      Visibility <- "504_Tank Grouping_DB2020_GROUP of TANK 3"
   Circle "Circle_23" at 1000,464 size 14x14
      Appearance <- "20_TANKS_IP_DATA_RIO_01_THIRD_TANK_BWT_LEVEL_HIHI"
   TextField "Text field_126" at 955,465 size 51x14; Text 'LS422-1S'
   Polyline "Polyline_7" at 921,458 size 123x259
      Visibility <- "504_Tank Grouping_DB2020_RUN TANK 3"
   TextField "Text field_10" at 950,618 size 74x20; Text 'Tank - 1S'
   Bar "Bar_9" at 790,459 size 122x258; MinimumValue 0; MaximumValue 100
      ProcessValue <- "20_TANKS_IP_DATA_RIO_02_FIRST_TANK_TANKS_PRESS"
   Button "Button_34" at 801,662 size 100x25; TextOff 'DISABLED'
      on Release: function_efd93a16("Tank 2S Status", 168, 315, -1, 0, 1)
      Visibility <- "504_Tank Grouping_DB2020_GROUP of TANK 5"
   Circle "Circle_22" at 868,465 size 14x14
      Appearance <- "20_TANKS_IP_DATA_RIO_02_SECOND_TANK_BWT_LEVEL_HIHI"
   TextField "Text field_127" at 823,466 size 51x14; Text 'LS422-2S'
   Polyline "Polyline_8" at 789,458 size 123x259
      Visibility <- "504_Tank Grouping_DB2020_RUN TANK 5"
   TextField "Text field_11" at 817,618 size 74x20; Text 'Tank - 2S'
   Bar "Bar_10" at 659,460 size 122x258; MinimumValue 0; MaximumValue 100
      ProcessValue <- "20_TANKS_IP_DATA_RIO_03_FIRST_TANK_TANKS_PRESS"
   Button "Button_38" at 669,663 size 100x25; TextOff 'DISABLED'
      on Release: function_efd93a16("Tank 3S Status", 168, 315, -1, 0, 1)
      Visibility <- "504_Tank Grouping_DB2020_GROUP of TANK 7"
   Circle "Circle_21" at 736,467 size 14x14
      Appearance <- "20_TANKS_IP_DATA_RIO_03_SECOND_TANK_BWT_LEVEL_HIHI"
   TextField "Text field_128" at 691,468 size 51x14; Text 'LS422-3S'
   Polyline "Polyline_9" at 658,458 size 123x259
      Visibility <- "504_Tank Grouping_DB2020_RUN TANK 7"
   TextField "Text field_12" at 690,618 size 74x20; Text 'Tank - 3S'
   Bar "Bar_11" at 526,459 size 122x258; MinimumValue 0; MaximumValue 100
      ProcessValue <- "20_TANKS_IP_DATA_RIO_04_FIRST_TANK_TANKS_PRESS"
   Button "Button_42" at 537,662 size 100x25; TextOff 'DISABLED'
      on Release: function_efd93a16("Tank 4S Status", 168, 315, -1, 2, 1)
      Visibility <- "504_Tank Grouping_DB2020_GROUP of TANK 9"
   Circle "Circle_19" at 604,466 size 14x14
      Appearance <- "20_TANKS_IP_DATA_RIO_04_SECOND_TANK_BWT_LEVEL_HIHI"
   TextField "Text field_129" at 559,467 size 51x14; Text 'LS422-4S'
   Polyline "Polyline_10" at 525,458 size 123x259
      Visibility <- "504_Tank Grouping_DB2020_RUN TANK 9"
   TextField "Text field_13" at 554,618 size 74x20; Text 'Tank - 4S'
   Bar "Bar_12" at 394,459 size 122x258; MinimumValue 0; MaximumValue 100
      ProcessValue <- "20_TANKS_IP_DATA_RIO_05_FIRST_TANK_TANKS_PRESS"
   Button "Button_46" at 405,662 size 100x25; TextOff 'DISABLED'
      on Release: function_efd93a16("Tank 5S Status", 168, 315, -1, 2, 1)
      Visibility <- "504_Tank Grouping_DB2020_GROUP of TANK 11"
   Circle "Circle_18" at 472,465 size 14x14
      Appearance <- "20_TANKS_IP_DATA_RIO_05_SECOND_TANK_BWT_LEVEL_HIHI"
   TextField "Text field_130" at 427,466 size 51x14; Text 'LS422-5S'
   Polyline "Polyline_11" at 393,458 size 123x259
      Visibility <- "504_Tank Grouping_DB2020_RUN TANK 11"
   TextField "Text field_18" at 424,618 size 74x20; Text 'Tank - 5S'
   Bar "Bar_13" at 262,460 size 122x258; MinimumValue 0; MaximumValue 100
      ProcessValue <- "20_TANKS_IP_DATA_RIO_06_FIRST_TANK_TANKS_PRESS"
   Button "Button_50" at 273,663 size 100x25; TextOff 'DISABLED'
      on Release: function_efd93a16("Tank 6S Status", 168, 315, -1, 2, 1)
      Visibility <- "504_Tank Grouping_DB2020_GROUP of TANK 13"
   Circle "Circle_17" at 340,467 size 14x14
      Appearance <- "20_TANKS_IP_DATA_RIO_06_SECOND_TANK_BWT_LEVEL_HIHI"
   TextField "Text field_131" at 295,468 size 51x14; Text 'LS422-6S'
   Polyline "Polyline_12" at 261,458 size 123x258
      Visibility <- "504_Tank Grouping_DB2020_RUN TANK 13"
   TextField "Text field_19" at 290,618 size 74x20; Text 'Tank - 6S'
   Bar "Bar_14" at 39,324 size 119x258; Unit %; MinimumValue 0; MaximumValue 100
      ProcessValue <- "20_TANKS_IP_DATA_RIO_07_FIRST_TANK_TANKS_PRESS"
   Circle "Circle_25" at 108,330 size 14x14
      Appearance <- "20_TANKS_IP_DATA_RIO_07_FIRST_TANK_BWT_LEVEL_HIHI"
   TextField "Text field_132" at 79,330 size 35x14; Text 'LS425'
   Polyline "Polyline_13" at 38,324 size 121x259
      Visibility <- "504_Tank Grouping_DB2020_RUN TANK 14"
   Button "Button_58" at 48,527 size 100x25; TextOff 'DISABLED'
      on Release: function_efd93a16("Tank AP Status", 168, 315, -1, 2, 1)
      Visibility <- "504_Tank Grouping_DB2020_GROUP of TANK 14"
   Button "HmiScreenItemData_6" at 1043,144 size 116x50; TextOn 'Back'; TextOff 'Tank Status'
      on Release: ActivateScreen("Balast Water Treatment Plant", 0)
   Button "Button_2" at 252,437 size 37x30; TextOff 'DB&B'
      on Release: function_efd93a16("Double Block & Bleed Valve Monitoring", 250, 250, -1, -1, 1)
      Appearance <- "10_DI_DATA_CV407_OPN"
   TextField "Text field_65" at 190,398 size 46x25; Text 'PGC'
   TextField "Text field_75" at 183,480 size 60x20; Text 'Disabled'
   TextField "Text field_76" at 183,480 size 60x20; Text 'Enabled'
      Visibility <- "10_DI_DATA_E_400_RUN"
   GraphicView "Graphic view_76" at 185,421 size 57x55; Picture "Graphic_251"
   Button "Button_6" at 179,402 size 70x105; TextOff 'Text'
      on Release: ActivateScreen("PGC System", 0)
   TextField "Text field_20" at 53,396 size 103x20; Text 'Aft PeakTank'
   GraphicView "Graphic view_108" at 4,683 size 96x48; Picture "Left Arow"
   Button "HmiScreenItemData_14" at 3,660 size 106x93; TextOn 'Back'; TextOff 'Text'
      on Press: ActivateScreen("Inert Gas Conditioning Plant", 0)
   IOField "I/O field_1" at 44,460 size 115x25; FormatPattern s999.9; Unit mBar
      ProcessValue <- "20_TANKS_IP_DATA_RIO_07_FIRST_TANK_TANKS_PRESS"
   IOField "I/O field_2" at 269,331 size 114x25; FormatPattern s999.9; Unit mBar
      ProcessValue <- "20_TANKS_IP_DATA_RIO_06_FIRST_TANK_TANKS_PRESS"
   IOField "I/O field_3" at 398,331 size 117x25; FormatPattern s999.9; Unit mBar
      ProcessValue <- "20_TANKS_IP_DATA_RIO_05_FIRST_TANK_TANKS_PRESS"
   IOField "I/O field_4" at 531,331 size 117x25; FormatPattern s999.9; Unit mBar
      ProcessValue <- "20_TANKS_IP_DATA_RIO_04_FIRST_TANK_TANKS_PRESS"
   IOField "I/O field_5" at 662,331 size 114x25; FormatPattern s999.9; Unit mBar
      ProcessValue <- "20_TANKS_IP_DATA_RIO_03_FIRST_TANK_TANKS_PRESS"
   IOField "I/O field_6" at 796,331 size 119x25; FormatPattern s999.9; Unit mBar
      ProcessValue <- "20_TANKS_IP_DATA_RIO_02_FIRST_TANK_TANKS_PRESS"
   IOField "I/O field_7" at 928,331 size 118x25; FormatPattern s999.9; Unit mBar
      ProcessValue <- "20_TANKS_IP_DATA_RIO_01_FIRST_TANK_TANKS_PRESS"
   IOField "I/O field_8" at 1103,459 size 119x25; FormatPattern s999.9; Unit mBar
      ProcessValue <- "20_TANKS_IP_DATA_RIO_01_FIRST_TANK_TANKS_PRESS"
   IOField "I/O field_9" at 928,555 size 118x25; FormatPattern s999.9; Unit mBar
      ProcessValue <- "20_TANKS_IP_DATA_RIO_01_FIRST_TANK_TANKS_PRESS"
   IOField "I/O field_10" at 796,556 size 118x25; FormatPattern s999.9; Unit mBar
      ProcessValue <- "20_TANKS_IP_DATA_RIO_02_FIRST_TANK_TANKS_PRESS"
   IOField "I/O field_11" at 664,558 size 116x25; FormatPattern s999.9; Unit mBar
      ProcessValue <- "20_TANKS_IP_DATA_RIO_03_FIRST_TANK_TANKS_PRESS"
   IOField "I/O field_12" at 530,557 size 117x25; FormatPattern s999.9; Unit mBar
      ProcessValue <- "20_TANKS_IP_DATA_RIO_04_FIRST_TANK_TANKS_PRESS"
   IOField "I/O field_13" at 400,558 size 114x25; FormatPattern s999.9; Unit mBar
      ProcessValue <- "20_TANKS_IP_DATA_RIO_05_FIRST_TANK_TANKS_PRESS"
   IOField "I/O field_14" at 268,559 size 116x25; FormatPattern s999.9; Unit mBar
      ProcessValue <- "20_TANKS_IP_DATA_RIO_06_FIRST_TANK_TANKS_PRESS"
   Button "Button_88" at 34,324 size 127x264; TextOff 'Text'
      on Release: function_efd93a16("Tank AP Status", 168, 315, -1, 0, 1)
      Appearance <- "504_Tank Grouping_DB2020_RUN TANK 14"
   Button "Button_86" at 259,458 size 126x260; TextOff 'Text'
      on Release: function_efd93a16("Tank 6S Status", 168, 315, -1, 0, 1)
      Appearance <- "504_Tank Grouping_DB2020_RUN TANK 13"
   Button "Button_79" at 391,457 size 126x262; TextOff 'Text'
      on Release: function_efd93a16("Tank 5S Status", 168, 315, -1, 0, 1)
      Appearance <- "504_Tank Grouping_DB2020_RUN TANK 11"
   Button "Button_77" at 523,457 size 126x262; TextOff 'Text'
      on Release: function_efd93a16("Tank 4S Status", 168, 315, -1, 0, 1)
      Appearance <- "504_Tank Grouping_DB2020_RUN TANK 9"
   Button "Button_74" at 657,457 size 126x262; TextOff 'Text'
      on Release: function_efd93a16("Tank 3S Status", 168, 315, -1, 0, 1)
      Appearance <- "504_Tank Grouping_DB2020_RUN TANK 7"
   Button "Button_70" at 788,457 size 126x262; TextOff 'Text'
      on Release: function_efd93a16("Tank 2S Status", 168, 315, -1, 0, 1)
      Appearance <- "504_Tank Grouping_DB2020_RUN TANK 5"
   Button "Button_66" at 921,457 size 126x261; TextOff 'Text'
      on Release: function_efd93a16("Tank 1S Status", 168, 315, -1, 0, 1)
      Appearance <- "504_Tank Grouping_DB2020_RUN TANK 3"
   Button "Button_61" at 1093,328 size 130x248; TextOff 'Text'
      on Release: function_efd93a16("Tank FP Status", 168, 315, -1, 0, 1)
      Appearance <- "504_Tank Grouping_DB2020_RUN TANK 1"
   Button "Button_62" at 919,205 size 126x242; TextOff 'Text'
      on Release: function_efd93a16("Tank 1P Status", 168, 315, -1, 0, 1)
      Appearance <- "504_Tank Grouping_DB2020_RUN TANK 2"
   Button "Button_68" at 789,202 size 126x246; TextOff 'Text'
      on Release: function_efd93a16("Tank 2P Status", 168, 315, -1, 0, 1)
      Appearance <- "504_Tank Grouping_DB2020_RUN TANK 4"
   Button "Button_72" at 654,205 size 126x242; TextOff 'Text'
      on Release: function_efd93a16("Tank 3P Status", 168, 315, -1, 0, 1)
      Appearance <- "504_Tank Grouping_DB2020_RUN TANK 6"
   Button "Button_76" at 524,205 size 126x243; TextOff 'Text'
      on Release: function_efd93a16("Tank 4P Status", 168, 315, -1, 0, 1)
      Appearance <- "504_Tank Grouping_DB2020_RUN TANK 8"
   Button "Button_78" at 392,206 size 126x241; TextOff 'Text'
      on Release: function_efd93a16("Tank 5P Status", 168, 315, -1, 0, 1)
      Appearance <- "504_Tank Grouping_DB2020_RUN TANK 10"
   Button "Button_84" at 259,204 size 126x244; TextOff 'Text'
      on Release: function_efd93a16("Tank 6P Status", 168, 315, -1, 0, 1)
      Appearance <- "504_Tank Grouping_DB2020_RUN TANK 12"
   Group "Group_5" at 664,46 size 45x27; FormatPattern 999
   Group "Group_1" at 711,46 size 50x27; FormatPattern 999; Unit h
   Group "Group_2" at 605,46 size 57x27; FormatPattern 999; Unit h
   Button "HmiScreenItemData_5" at 180,144 size 116x50; TextOn 'Back'; TextOff 'Tank Status'
      on Release: function_efd93a16("Tank Status", 400, 250, -1, -1, 1)
   Button "Button_10" at 14,93 size 153x55; TextOff 'Text'
      on Release: function_efd93a16("Salinity - Acceptance", 168, 315, -1, 0, 1)
      Visibility <- "2068_Sys_Status_Data_SAL_VALID"
   Button "Button_12" at 14,93 size 153x53; TextOff 'Text'
      on Release: function_efd93a16("Tank Times", 300, 200, -1, 0, 1)
      Visibility <- "2068_Sys_Status_Data_Times Visibil"
   Button "Button_59" at 298,44 size 240x30; TextOn 'TB3 Enabled'; TextOff 'BWT System Shutting Down'
      Visibility <- "2110_BTCS_CNTRL_DB_BTCS_STATE"
   Button "Button_60" at 299,44 size 240x30; TextOn 'TB3 Enabled'; TextOff 'BWT System Enabled'
      Visibility <- "2110_BTCS_CNTRL_DB_BTCS_STATE"
   IOField "I/O field_29" at 664,46 size 45x27; FormatPattern 99; Unit h
      ProcessValue <- "Sequence Times_DB_Treatment Timer_Hours Left"
      Visibility <- "2110_BTCS_CNTRL_DB_BTCS_STATE"
   IOField "I/O field_30" at 664,46 size 45x27; FormatPattern 99; Unit h
      ProcessValue <- "Sequence Times_DB_Pre-Dwell Timer_Hours Left"
      Visibility <- "2110_BTCS_CNTRL_DB_BTCS_STATE"
   IOField "I/O field_15" at 711,46 size 50x27; FormatPattern 99; Unit m
      ProcessValue <- "Sequence Times_DB_Treatment Timer_Minutes Left"
      Visibility <- "2110_BTCS_CNTRL_DB_BTCS_STATE"
   IOField "I/O field_16" at 711,46 size 50x27; FormatPattern 99; Unit m
      ProcessValue <- "Sequence Times_DB_Pre-Dwell Timer_Minutes Left"
      Visibility <- "2110_BTCS_CNTRL_DB_BTCS_STATE"
   IOField "I/O field_17" at 605,46 size 57x27; FormatPattern 999; Unit d
      ProcessValue <- "Sequence Times_DB_Treatment Timer_Days Left"
      Visibility <- "2110_BTCS_CNTRL_DB_BTCS_STATE"
   IOField "I/O field_18" at 605,46 size 57x27; FormatPattern 999; Unit d
      ProcessValue <- "Sequence Times_DB_Pre-Dwell Timer_Days Left"
      Visibility <- "2110_BTCS_CNTRL_DB_BTCS_STATE"

VB script "VoyageTimeInsufficient"
   If SmartTags("Voyage Time Invalid") Then
   	efd93a16-2665-4b85-bcb9-25eddcb7b6f4 Voyage Time Warning,275,250,$3$hmiOn$,$3$hmiTop$,$3$hmiMedium$
   ElseIf Not SmartTags("Voyage Time Invalid") Then
   	efd93a16-2665-4b85-bcb9-25eddcb7b6f4Voyage Time Warning,0,0,$3$hmiOff$,$3$hmiAnimationOff$,$3$hmiMedium$
   End If

VB script "TreatmentCycleCompleted"
   If SmartTags("Sequence Times_DB_Post-Dwell Timer_Q") Then
   	efd93a16-2665-4b85-bcb9-25eddcb7b6f4 Treatment Cycle Completed,275,250,$3$hmiOn$,$3$hmiBottom$,$3$hmiMedium$
   'ElseIf Not SmartTags("Treatment Runs Completed") Then
   '	ShowPopupScreen"Treatment Cycle Completed",0,0,hmiOff,hmiAnimationOff,hmiMedium
   End If

VB script "SD_Card_Overflow"
   If SmartTags("Logging SD Card Overflow") Then 
   	efd93a16-2665-4b85-bcb9-25eddcb7b6f4 SD Card overflow,275,250,$3$hmiOn$,$3$hmiBottom$,$3$hmiMedium$
   ElseIf Not SmartTags("Logging SD Card Overflow") Then
   	efd93a16-2665-4b85-bcb9-25eddcb7b6f4SD Card overflow,0,0,$3$hmiOff$,$3$hmiAnimationOff$,$3$hmiMedium$
   End If

VB script "Salinity_FreshWaterAlert"
   If SmartTags("2068_Sys_Status_Data_SAL_CNF_CHK") Then
   	efd93a16-2665-4b85-bcb9-25eddcb7b6f4 Salinity - Fresh Water Alert,789,316,$3$hmiOn$,$3$hmiBottom$,$3$hmiMedium$
   ElseIf Not SmartTags("2068_Sys_Status_Data_SAL_CNF_CHK") Then
   	efd93a16-2665-4b85-bcb9-25eddcb7b6f4Salinity - Fresh Water Alert,0,0,$3$hmiOff$,$3$hmiAnimationOff$,$3$hmiMedium$
   End If

VB script "TimeRemainingToTreatment"
   If SmartTags("Warn To Start IGG") Then
   	efd93a16-2665-4b85-bcb9-25eddcb7b6f4 Time Until Treatment Required, 400, 200, $3$hmiOn$, $3$hmiBottom$, $3$hmiMedium$
   	ElseIf Not SmartTags("Warn To Start IGG") Then
   efd93a16-2665-4b85-bcb9-25eddcb7b6f4 Time Until Treatment Required, 0, 0, $3$hmiOff$, $3$hmiOff$, $3$hmiMedium$
   End If

VB script "TreatmentRequired"
   If SmartTags("Warn To Start IGG-Last") Then
   	efd93a16-2665-4b85-bcb9-25eddcb7b6f4 Start Treatment, 400, 200, $3$hmiOn$, $3$hmiBottom$, $3$hmiMedium$
   	ElseIf Not SmartTags("Warn To Start IGG-Last") Then
   efd93a16-2665-4b85-bcb9-25eddcb7b6f4 Start Treatment, 0, 0, $3$hmiOff$, $3$hmiOff$, $3$hmiMedium$
   End If

VB script "PGCCommissioning"
   If SmartTags("PGC_COMMISSION_MODE_DB_Drive Popup") Then
   	efd93a16-2665-4b85-bcb9-25eddcb7b6f4 PGC Commissioning, 0, 0, $3$hmiOn$, $3$hmiBottom$, $3$hmiMedium$
   	ElseIf Not SmartTags("PGC_COMMISSION_MODE_DB_Drive Popup") Then
   efd93a16-2665-4b85-bcb9-25eddcb7b6f4 PGC Commissioning, 0, 0, $3$hmiOff$, $3$hmiOff$, $3$hmiMedium$
   End If

VB script "User_Change"
   f41c6f6c-971d-4734-9362-16d81ac70597 Current User
   e1ab61de-e5a2-437b-97c4-abda991a3a2e user_group
   
   'Tip:
   ' 1. Use the <CTRL+SPACE> or <CTRL+I> shortcut to open a list of all objects and functions
   ' 2. Write the code using the HMI Runtime object.
   '  Example: HmiRuntime.Screens("Screen_1").
   ' 3. Use the <CTRL+J> shortcut to create an object reference.
   'Write the code as of this position:

VB script "TreatmentdDailyChecks"
   If SmartTags("88_treatment_POP_UP") Then
   	efd93a16-2665-4b85-bcb9-25eddcb7b6f4 Treatment check / Daily Checks Completed,275,250,$3$hmiOn$,$3$hmiBottom$,$3$hmiMedium$
   End If

VB script "TitleUpdater"
   Dim title
   Set title = HmiRuntime.ActiveScreen.ScreenItems("Screen title")
   title.Text = HmiRuntime.ActiveScreen.ObjectName

VB script "BWT_Warning"
   If SmartTags("2068_Sys_Status_Data_Not BWT mode Warning") Then
   	efd93a16-2665-4b85-bcb9-25eddcb7b6f4 BWT Mode Warning,275,250,$3$hmiOn$,$3$hmiTop$,$3$hmiMedium$
   'ElseIf Not SmartTags("BWT Mode Warning") Then
   '	ShowPopupScreen"BWT Mode Warning",0,0,hmiOff,hmiAnimationOff,hmiMedium
   End If

VB script "Report_Test"
   f41c6f6c-971d-4734-9362-16d81ac70597 Current User
   e1ab61de-e5a2-437b-97c4-abda991a3a2e user_group
   
   
   'Tip:
   ' 1. Use the <CTRL+SPACE> or <CTRL+I> shortcut to open a list of all objects and functions
   ' 2. Write the code using the HMI Runtime object.
   '  Example: HmiRuntime.Screens("Screen_1").
   ' 3. Use the <CTRL+J> shortcut to create an object reference.
   'Write the code as of this position:

VB script "HeartBeatFunction"
   If SmartTags("IGG HMI HEART BEAT")=0 Then
   	b21d3eaf-4e31-425c-ad1a-ba4e4002cacc(IGG HMI HEART BEAT),1
   Else
   	b21d3eaf-4e31-425c-ad1a-ba4e4002cacc (IGG HMI HEART BEAT),0
   End If

VB script "HeartBeatHMI_Warning"
   Dim Warning, Tempos
   
   
   If SmartTags("HEART BEAT TRUE")=True Then
   	Warning=0 '"HEART BEAT TRUE"
   Else
   	Warning=1
   End If
   
   If Warning=0 Then
   	efd93a16-2665-4b85-bcb9-25eddcb7b6f4 Lost Comunication, 0, 0, $3$hmiOff$, $3$hmiOff$, $3$hmiMedium$
   Else
   	efd93a16-2665-4b85-bcb9-25eddcb7b6f4 Lost Comunication, 300, 100, $3$hmiOn$, $3$hmiBottom$, $3$hmiMedium$
   End If		
   
   	b21d3eaf-4e31-425c-ad1a-ba4e4002cacc SmartTags("HEART BEAT TRUE"),False

VB script "PGC_ProtectionWarning"
   If SmartTags("Setpoint Override_DB_Set Pressure") Then
   	efd93a16-2665-4b85-bcb9-25eddcb7b6f4 PGC Protection Warning,275,250,$3$hmiOn$,$3$hmiTop$,$3$hmiMedium$
   'ElseIf Not SmartTags("Setpoint Override_DB_Set Pressure") Then
   '	ShowPopupScreen"Setpoint Override_DB_Set Pressure",0,0,hmiOff,hmiAnimationOff,hmiMedium
   End If

VB script "ALARM_Present"
   If SmartTags("60_Alarm_Data_ALRM_PRSNT") Then
   	bec8f1e5-2ab1-45f6-ad91-1d37c469eb91 04 Alarm Log,0
   End If
   
   'If Not SmartTags("60_Alarm_Data_ALRM_PRSNT") Then
   '	ActivateScreen "01 Home",0
   'End If
   
   
   
   
   
   
   
   
   
   'Tip:
   ' 1. Use the <CTRL+SPACE> or <CTRL+I> shortcut to open a list of all objects and functions
   ' 2. Write the code using the HMI Runtime object.
   '  Example: HmiRuntime.Screens("Screen_1").
   ' 3. Use the <CTRL+J> shortcut to create an object reference.
   'Write the code as of this position:

VB script "TreatmentRequired_GCU"
   If SmartTags("Warn To Start GCU-Last") Then
   	efd93a16-2665-4b85-bcb9-25eddcb7b6f4 Start GCU for Re-Ox, 400, 200, $3$hmiOn$, $3$hmiBottom$, $3$hmiMedium$
   	ElseIf Not SmartTags("Warn To Start GCU-Last") Then
   efd93a16-2665-4b85-bcb9-25eddcb7b6f4 Start GCU for Re-Ox, 0, 0, $3$hmiOff$, $3$hmiOff$, $3$hmiMedium$
   End If

VB script "TimeRemainingToRe_Ox"
   If SmartTags("Warn To Start GCU") Then
   	efd93a16-2665-4b85-bcb9-25eddcb7b6f4 Time Until GCU Start Required, 400, 200, $3$hmiOn$, $3$hmiBottom$, $3$hmiMedium$
   	ElseIf Not SmartTags("Warn To Start GCU") Then
   efd93a16-2665-4b85-bcb9-25eddcb7b6f4 Time Until GCU Start Required, 0, 0, $3$hmiOff$, $3$hmiOff$, $3$hmiMedium$
   End If

VB script "TANK_Activ_Warning"
   If SmartTags("Not TANK Activ Warning") Then
   	efd93a16-2665-4b85-bcb9-25eddcb7b6f4 TANK Activ Warning,300,200,$3$hmiOn$,$3$hmiTop$,$3$hmiMedium$
   'ElseIf Not SmartTags("Not TANK Activ Warning") Then
   '	ShowPopupScreen"TANK Activ Warning",0,0,hmiOff,hmiAnimationOff,hmiMedium
   End If

scheduled task "VB procces"
   Triggers <- "1 min"

scheduled task "User Change"
   on Action: "User_Change"()

scheduled task "Heart Beat"
   on Action: "HeartBeatFunction"(); "HeartBeatHMI_Warning"()
   Triggers <- "1 min"
*)

(* ===== HMI "HMI_RT_4" =====
system functions are stored by id; their names below are inferred from use
connection "IGG PLC Comms_3": ETHERNET, S7_1500_OMS
connection "BC PLC Comms_3": ETHERNET, S7_1500_OMS
connection "BWTS PLC Comms_3": ETHERNET, S7_1500_OMS

HMI tags "Default tag table"
   "66_Event_Data_BC_EVENT_WORD_01" : Word = PLC "66_Event_Data".BC_EVENT_WORD_01 AT %DB66.DBW0, 1 s
   "66_Event_Data_BC_EVENT_WORD_02" : Word = PLC "66_Event_Data".BC_EVENT_WORD_02 AT %DB66.DBW2, 1 s
   "64_Message_Data_BC_MESSAGE_WORD_01" : Word = PLC "64_Message_Data".BC_MESSAGE_WORD_01 AT %DB64.DBW0, 1 s
   "64_Message_Data_BC_MESSAGE_WORD_02" : Word = PLC "64_Message_Data".BC_MESSAGE_WORD_02 AT %DB64.DBW2, 1 s
   "66_Event_Data_IGG_EVENT_WORD_01" : Word = PLC "66_Event_Data".IGG_EVENT_WORD_01 AT %DB66.DBW0, 1 s
   "66_Event_Data_IGG_EVENT_WORD_02" : Word = PLC "66_Event_Data".IGG_EVENT_WORD_02 AT %DB66.DBW2, 1 s
   "64_Message_Data_IGG_MESSAGE_WORD_01" : Word = PLC "64_Message_Data".IGG_MESSAGE_WORD_01 AT %DB64.DBW0, 1 s
   "64_Message_Data_IGG_MESSAGE_WORD_02" : Word = PLC "64_Message_Data".IGG_MESSAGE_WORD_02 AT %DB64.DBW2, 1 s
   "Current User" : WString[15] AT %DB1.DBX0.0
   "db_time_sync_time_system_READ" : LDT = PLC db_time_sync_time_system_READ AT %M2.0, 1 s
   "80_From_HMI_Cooling System Overrun" : Time = PLC "80_From_HMI"."Cooling System Overrun", 1 s
   "db_time_sync_time_local_READ" : LDT = PLC db_time_sync_time_local_READ AT %M4.0, 1 s
   "82_To_HMI_Fuel Pump 1 Animation" : Int = PLC "82_To_HMI"."Fuel Pump 1 Animation", 1 s
   "82_To_HMI_Fuel Pump 2 Animation" : Int = PLC "82_To_HMI"."Fuel Pump 2 Animation", 1 s
   "16_AQ_Data_CV203_CNTRL(1)" : Real = PLC "16_AQ_Data".CV203_CNTRL, 1 s
   "HMI Data_O2 Setpoint" : Real, internal
   "82_To_HMI_IA Compressor Animation" : Int = PLC "82_To_HMI"."IA Compressor Animation", 1 s
   "Atomising Air  Valve Manual Regulator" : Int, internal
   "Fuel Valve Manual Regulator" : Int, internal
   "82_To_HMI_I&A Compressor Run Hours(1)" : Int = PLC "82_To_HMI"."I&A Compressor Run Hours", 1 s
   "82_To_HMI_I&A Compressor Service Time Hours" : Int = PLC "82_To_HMI"."I&A Compressor Service Time Hours", 1 s
   "82_To_HMI_CA Blower Run Days" : Int = PLC "82_To_HMI"."CA Blower Run Days", 1 s
   "82_To_HMI_CA Blower Service Time Hours" : Int = PLC "82_To_HMI"."CA Blower Service Time Hours", 1 s
   "82_To_HMI_CA Blower Run Hours" : Int = PLC "82_To_HMI"."CA Blower Run Hours", 1 s
   "82_To_HMI_CA Blower Run Minutes" : Int = PLC "82_To_HMI"."CA Blower Run Minutes", 1 s
   "82_To_HMI_I&A Compressor Run Minutes" : Int = PLC "82_To_HMI"."I&A Compressor Run Minutes", 1 s
   "82_To_HMI_I&A Compressor Run Seconds" : Int = PLC "82_To_HMI"."I&A Compressor Run Seconds", 1 s
   "P305_Functioning Hours_IDB_Hours Total" : Int = PLC "P305_Functioning Hours_IDB"."Hours Total", 1 s
   "HMI Data_Fresh Water Service Time" : Int, internal
   "P305_Functioning Hours_IDB_Service Time bit" : Bool = PLC "P305_Functioning Hours_IDB"."Service Time bit", 1 s
   "P305_Functioning Hours_IDB_Minutes" : Int = PLC "P305_Functioning Hours_IDB".Minutes, 1 s
   "P305_Functioning Hours_IDB_Seconds" : Int = PLC "20_TANKS_IP_DATA".RIO_04.SECOND_TANK.BWT_LEVEL_HIHI, 1 s
   "FW Pump Animation" : Int, internal
   "82_To_HMI_I&A Compressor Run Hours" : Int = PLC "82_To_HMI"."I&A Compressor Run Hours", 1 s
   "82_To_HMI_CRNT_MODE_IGG" : Int = PLC "82_To_HMI".CRNT_MODE_IGG, 1 s
   "70_Mode_Data_AUT_RST_PLS_IN" : Bool = PLC "70_Mode_Data".AUT_RST_PLS.IN, 1 s
   "100_IGG_AUTO_SEQ_DB_CRNT_STEP" : Int = PLC "100_IGG_AUTO_SEQ_DB".CRNT_STEP, 1 s
   "100_BC_AUTO_SEQ_DB_CRNT_STEP" : Int = PLC "100_BC_AUTO_SEQ_DB".CRNT_STEP, 1 s
   "103_Main_Burner_DB_RUN" : Bool = PLC "103_Main_Burner_DB".RUN, 1 s
   "60_Alarm_Data_ALRM_PRSNT" : Bool = PLC "60_Alarm_Data".ALRM_PRSNT AT %DB60.DBX32.0, 1 s
      on ChangeValue: "ALARM_Present"()
   "62_Warning_Data_WRNG_PRSNT" : Bool = PLC "62_Warning_Data".WRNG_PRSNT AT %DB62.DBX16.0, 1 s
   "103_Main_Burner_DB_RUNNING" : Bool = PLC "103_Main_Burner_DB".RUNNING, 1 s
   "101_Fuel_Pumps_DB_Duty Is B" : Bool = PLC "101_Fuel_Pumps_DB"."Duty Is B", 1 s
   "101_Fuel_Pumps_DB_Duty Is A" : Bool = PLC "101_Fuel_Pumps_DB"."Duty Is A", 1 s
   "84_Setpoints_PIT204_High" : Real = PLC "84_Setpoints".PIT204_High, 1 s
   "84_Setpoints_PIT204_High(1)" : Real = PLC "84_Setpoints".PIT204_High, 1 s
   "84_Setpoints_PIT204_HighHigh" : Real = PLC "84_Setpoints".PIT204_HighHigh, 1 s
   "84_Setpoints_PIT204_HighHigh(1)" : Real = PLC "84_Setpoints".PIT204_HighHigh, 1 s
   "84_Setpoints_PIT204_LowLow" : Real = PLC "84_Setpoints".PIT204_LowLow, 1 s
   "84_Setpoints_PIT204_LowLow(1)" : Real = PLC "84_Setpoints".PIT204_LowLow, 1 s
   "84_Setpoints_PIT204_Low" : Real = PLC "84_Setpoints".PIT204_Low, 1 s
   "84_Setpoints_PIT204_Low(1)" : Real = PLC "84_Setpoints".PIT204_Low, 1 s
   "80_From_HMI_RST_LOCKOUT" : Bool = PLC "80_From_HMI".RST_LOCKOUT, 1 s
   "80_From_HMI_Beacon frequency" : Time = PLC "80_From_HMI"."Beacon frequency", 1 s
   "80_From_HMI_Buzzer reset time" : Time = PLC "80_From_HMI"."Buzzer reset time", 1 s
   "80_From_HMI_Reset_Alarms" : Bool = PLC "80_From_HMI".Reset_Alarms, 1 s
   "Alarm beacon handling_DB_Buzzer_Timer_0_Instance_Q" : Bool = PLC "Alarm beacon handling_DB".Buzzer_Timer_0_Instance.Q, 1 s
   "Buzzer" : Bool = PLC Buzzer AT %Q1.7, 1 s
   "80_From_HMI_FLM_FAIL_DLY" : Time = PLC "80_From_HMI".FLM_FAIL_DLY, 1 s
   "103_Main_Burner_DB_DN_OK" : Bool = PLC "103_Main_Burner_DB".DN_OK, 1 s
   "103_Main_Burner_DB_Days burn_CV" : Int = PLC "103_Main_Burner_DB"."Days burn".CV, 1 s
   "103_Main_Burner_DB_Hours burn_CV" : Int = PLC "103_Main_Burner_DB"."Hours burn".CV, 1 s
   "103_Main_Burner_DB_Minutes burn_CV" : Int = PLC "103_Main_Burner_DB"."Minutes burn".CV, 1 s
   "103_Main_Burner_DB_Seconds burn_CV" : Int = PLC "103_Main_Burner_DB"."Seconds burn".CV, 1 s
   "103_Main_Burner_DB_STATE" : Int = PLC "103_Main_Burner_DB".STATE, 1 s
   "19_AUTO_CMNDS_Data_CV203_RAMP_CNTRL" : Bool = PLC "19_AUTO_CMNDS_Data".CV203_RAMP_CNTRL, 1 s
   "102_Pilot_Burner_DB_RUNNING" : Bool = PLC "102_Pilot_Burner_DB".RUNNING, 1 s
   "68_Sys_Status_Data_FUEL_PRES_IN_RNG" : Bool = PLC "68_Sys_Status_Data".FUEL_PRES_IN_RNG, 1 s
   "68_Sys_Status_Data_IA_PRES_IN_RNG" : Bool = PLC "68_Sys_Status_Data".IA_PRES_IN_RNG, 1 s
   "84_Setpoints_Gain" : Real = PLC "84_Setpoints".Gain, 1 s
   "84_Setpoints_Integration Time" : Time = PLC "84_Setpoints"."Integration Time", 1 s
   "84_Setpoints_Derive Time" : Time = PLC "84_Setpoints"."Derive Time", 1 s
   "O2 Ramp Control_QLMN_HLM" : Bool = PLC "O2 Ramp Control".QLMN_HLM, 1 s
   "O2 Ramp Control_QLMN_LLM" : Bool = PLC "O2 Ramp Control".QLMN_LLM, 1 s
   "84_Setpoints_P_ON" : Bool = PLC "84_Setpoints".P_ON, 1 s
   "84_Setpoints_I_ON" : Bool = PLC "84_Setpoints".I_ON, 1 s
   "84_Setpoints_D_ON" : Bool = PLC "84_Setpoints".D_ON, 1 s
   "Evolving Setpoint_DB_LevelBetter" : Bool = PLC "Evolving Setpoint_DB".LevelBetter, 1 s
   "84_Setpoints_Max Opening" : Real = PLC "84_Setpoints"."Max Opening", 1 s
   "84_Setpoints_Min Opening" : Real = PLC "86_Times".STEP_MAX_TIME_STP_290, 1 s
   "80_From_HMI_Post Purge Time" : Time = PLC "80_From_HMI"."Post Purge Time", 1 s
   "103_Main_Burner_DB_Status" : Int = PLC "103_Main_Burner_DB".Status, 1 s
   "80_From_HMI_Reset CV203 PID" : Bool = PLC "80_From_HMI"."Reset CV203 PID", 1 s
   "80_From_HMI_BurnerProgramedStop" : Bool = PLC "80_From_HMI".BurnerProgramedStop, 1 s
   "82_To_HMI_CA Blower Reset Hours" : Bool = PLC "82_To_HMI"."CA Blower Reset Hours", 1 s
   "82_To_HMI_CA Blower Service Due" : Bool = PLC "82_To_HMI"."CA Blower Service Due", 1 s
   "Operation hours E139_IDB_Hours Functioning" : Int = PLC "Operation hours E139_IDB"."Hours Functioning", 1 s
   "82_To_HMI_CA Blower Total Run Hours" : Int = PLC "82_To_HMI"."CA Blower Total Run Hours", 1 s
   "82_To_HMI_I&A Compressor Total Run Hours" : Int = PLC "82_To_HMI"."I&A Compressor Total Run Hours", 1 s
   "82_To_HMI_I&A Compressor Reset Hours" : Bool = PLC "82_To_HMI"."I&A Compressor Reset Hours", 1 s
   "82_To_HMI_I&A Compressor Service Due" : Bool = PLC "82_To_HMI"."I&A Compressor Service Due", 1 s
   "82_To_HMI_E500A Fuel Pump Run Hours" : Int = PLC "82_To_HMI"."E500A Fuel Pump Run Hours", 1 s
   "64_Functioning Hours_E500A_IDB_Hours Functioning" : Int = PLC "64_Functioning Hours_E500A_IDB"."Hours Functioning", 1 s
   "82_To_HMI_E500A Fuel Pump Run Minutes" : Int = PLC "82_To_HMI"."E500A Fuel Pump Run Minutes", 1 s
   "82_To_HMI_E500A Fuel Pump Run Seconds" : Int = PLC "82_To_HMI"."E500A Fuel Pump Run Seconds", 1 s
   "82_To_HMI_E500A Fuel Pump Total Run Hours" : Int = PLC "82_To_HMI"."E500A Fuel Pump Total Run Hours", 1 s
   "82_To_HMI_E500A Fuel Pump Service Time Hours" : Int = PLC "82_To_HMI"."E500A Fuel Pump Service Time Hours", 1 s
   "82_To_HMI_E500A Fuel Pump Reset Hours" : Bool = PLC "82_To_HMI"."E500A Fuel Pump Reset Hours", 1 s
   "64_Functioning Hours_E500B_IDB_Hours Functioning" : Int = PLC "64_Functioning Hours_E500B_IDB"."Hours Functioning", 1 s
   "82_To_HMI_E500B Fuel Pump Run Minutes" : Int = PLC "82_To_HMI"."E500B Fuel Pump Run Minutes", 1 s
   "82_To_HMI_E500B Fuel Pump Run Seconds" : Int = PLC "82_To_HMI"."E500B Fuel Pump Run Seconds", 1 s
   "82_To_HMI_E500B Fuel Pump Total Run Hours" : Int = PLC "82_To_HMI"."E500B Fuel Pump Total Run Hours", 1 s
   "82_To_HMI_E500B Fuel Pump Service Time Hours" : Int = PLC "82_To_HMI"."E500B Fuel Pump Service Time Hours", 1 s
   "82_To_HMI_E500B Fuel Pump Reset Hours" : Bool = PLC "82_To_HMI"."E500B Fuel Pump Reset Hours", 1 s
   "82_To_HMI_E500B Fuel Pump Service Due" : Bool = PLC "82_To_HMI"."E500B Fuel Pump Service Due", 1 s
   "82_To_HMI_E500A Fuel Pump Service Due" : Bool = PLC "82_To_HMI"."E500A Fuel Pump Service Due", 1 s
   "64_Functioning Hours_P301_IDB_Hours Functioning" : Int = PLC "64_Functioning Hours_P301_IDB"."Hours Functioning", 1 s
   "82_To_HMI_P301 CSW Pump Run Minutes" : Int = PLC "82_To_HMI"."P301 CSW Pump Run Minutes", 1 s
   "82_To_HMI_P301 CSW Pump Run Seconds" : Int = PLC "82_To_HMI"."P301 CSW Pump Run Seconds", 1 s
   "82_To_HMI_P301 CSW Pump Reset Hours" : Bool = PLC "82_To_HMI"."P301 CSW Pump Reset Hours", 1 s
   "82_To_HMI_P301 CSW Pump Service Due" : Bool = PLC "82_To_HMI"."P301 CSW Pump Service Due", 1 s
   "80_From_HMI_P301_PRSNT" : Bool = PLC "80_From_HMI".P301_PRSNT, 1 s
   "Alarms_Acknowledge_IGG_ALARM_ACKNLG_3" : Word = PLC Alarms_Acknowledge.IGG_ALARM_ACKNLG_3 AT %DB67.DBW4, 1 s
   "Alarms_Acknowledge_IGG_ALARM_ACKNLG_4" : Word = PLC Alarms_Acknowledge.IGG_ALARM_ACKNLG_4 AT %DB67.DBW6, 1 s
   "Alarms_Acknowledge_IGG_ALARM_ACKNLG_2" : Word = PLC Alarms_Acknowledge.IGG_ALARM_ACKNLG_2 AT %DB67.DBW2, 1 s
   "Alarms_Acknowledge_IGG_ALARM_ACKNLG_1" : Word = PLC Alarms_Acknowledge.IGG_ALARM_ACKNLG_1 AT %DB67.DBW0, 1 s
   "BC_ALARM_ACKNLG_1" : Word = PLC BC_ALARM_ACKNLG_1 AT %MW24, 1 s
   "BC_ALARM_ACKNLG_2" : Word = PLC BC_ALARM_ACKNLG_2 AT %MW26, 1 s
   "BC_ALARM_ACKNLG_3" : Word = PLC BC_ALARM_ACKNLG_3 AT %MW28, 1 s
   "BC_ALARM_ACKNLG_4" : Word = PLC BC_ALARM_ACKNLG_4 AT %MW30, 1 s
   "80_From_HMI_P305_PRSNT" : Bool = PLC "80_From_HMI".P305_PRSNT, 1 s
   "68_Sys_Status_Data_INTRLKS_OK" : Bool = PLC "68_Sys_Status_Data".INTRLKS_OK, 1 s
   "82_To_HMI_E-STOP LATCHED" : Bool = PLC "82_To_HMI"."E-STOP LATCHED", 1 s
   "82_To_HMI_P301 CSW Pump Run Days" : Int = PLC "82_To_HMI"."P301 CSW Pump Run Days", 1 s
   "82_To_HMI_CA Blower Run Seconds" : Int = PLC "82_To_HMI"."CA Blower Run Seconds", 1 s
   "82_To_HMI_P305 FW Pump Reset Hours" : Bool = PLC "82_To_HMI"."P305 FW Pump Reset Hours", 1 s
   "P305_Functioning Hours_IDB_Hours Functioning Out" : Int = PLC "P305_Functioning Hours_IDB"."Hours Functioning Out", 1 s
   "82_To_HMI_P305 FW Pump Run Hours" : Int = PLC "82_To_HMI"."P305 FW Pump Run Hours", 1 s
   "82_To_HMI_P305 FW Pump Run Days" : Int = PLC "82_To_HMI"."P305 FW Pump Run Days", 1 s
   "82_To_HMI_P301 CSW Pump Service Time Hours" : Int = PLC "82_To_HMI"."P301 CSW Pump Service Time Hours", 1 s
   "82_To_HMI_P301 CSW Pump Run Hours" : Int = PLC "82_To_HMI"."P301 CSW Pump Run Hours", 1 s
   "82_To_HMI_P301 CSW Pump Total Run Hours" : Int = PLC "82_To_HMI"."P301 CSW Pump Total Run Hours", 1 s
   "80_From_HMI_PIT 359 delay" : Time = PLC "80_From_HMI"."PIT 359 delay", 1 s
   "80_From_HMI_PIT 316 delay" : Time = PLC "80_From_HMI"."PIT 316 delay", 1 s
   "86_Times_PIT402_Ramp_Seconds" : Int = PLC "86_Times".PIT402_Ramp_Seconds, 1 s
   "86_Times_PIT402 Alarm Delay" : Time = PLC "86_Times"."PIT402 Alarm Delay", 1 s
   "84_Setpoints_PIT113_Burner_Target" : Real = PLC "84_Setpoints".PIT113_Burner_Target, 1 s
   "1111_PID_CV111_Setpoint" : Real = PLC "1111_PID_CV111".Setpoint, 1 s
   "2062_Warning_Data_BTCS_WARNING_WORD_12" : Word = PLC "2062_Warning_Data".BTCS_WARNING_WORD_12 AT %DB2062.DBW362, 1 s
   "2062_Warning_Data_BTCS_WARNING_WORD_13" : Word = PLC "2062_Warning_Data".BTCS_WARNING_WORD_13 AT %DB2062.DBW364, 1 s
   "2062_Warning_Data_BTCS_WARNING_WORD_14" : Word = PLC "2062_Warning_Data".BTCS_WARNING_WORD_14 AT %DB2062.DBW366, 1 s
   "2062_Warning_Data_BTCS_WARNING_WORD_15" : Word = PLC "2062_Warning_Data".BTCS_WARNING_WORD_15 AT %DB2062.DBW368, 1 s
   "2062_Warning_Data_BTCS_WARNING_WORD_16" : Word = PLC "2062_Warning_Data".BTCS_WARNING_WORD_16 AT %DB2062.DBW370, 1 s
   "12_AI_Data_PIT113In_SCALED" : Real = PLC "12_AI_Data".PIT113In_SCALED, 1 s
   "PGC Flush_DB_PGC Stop Delay" : Time = PLC "PGC Flush_DB"."PGC Stop Delay", 1 s
   "PGC Flush_DB_CAB after Start Delay" : Time = PLC "PGC Flush_DB"."CAB after Start Delay", 1 s
   "PGC Flush_DB_CAB RPM Cmnd" : Real = PLC "PGC Flush_DB"."CAB RPM Cmd", 1 s
   "PGC Flush_DB_Override" : Bool = PLC "PGC Flush_DB".Override, 1 s
   "PGC Flush_DB_Running" : Bool = PLC "PGC Flush_DB".Running, 1 s
   "PGC Flush_DB_Activate" : Bool = PLC "PGC Flush_DB".Activate, 1 s
   "PGC Flush_DB_Done" : Bool = PLC "PGC Flush_DB".Done, 1 s
   "PGC Flush_DB_CV405 Open" : Bool = PLC "PGC Flush_DB"."CV405 Open", 1 s
   "PGC Flush_DB_CV401 Open" : Bool = PLC "PGC Flush_DB"."CV401 Open", 1 s
   "PGC Flush_DB_CV431 Open" : Bool = PLC "PGC Flush_DB"."CV431 Open", 1 s
   "PGC Flush_DB_CAB Start" : Bool = PLC "PGC Flush_DB"."CAB Start", 1 s
   "PGC Flush_DB_CV403 Modulate" : Bool = PLC "PGC Flush_DB"."CV403 Modulate", 1 s
   "PGC Flush_DB_Stop PGC" : Bool = PLC "PGC Flush_DB"."Stop PGC", 1 s
   "PGC Flush_DB_PGC Purge Duration" : Time = PLC "PGC Flush_DB"."PGC Purge Duration", 1 s
   "PGC Flush_DB_CV403 Open" : Bool = PLC "PGC Flush_DB"."CV403 Open", 1 s
   "PGC Flush_DB_Flip Flop_Override_Output" : Bool = PLC "PGC Flush_DB"."Flip Flop_Override".Output, 1 s
   "19_AUTO_CMNDS_Data_Purge Rqst Simulate" : Bool = PLC "19_AUTO_CMNDS_Data"."Purge Rqst Simulate", 1 s
   "PGC Flush_DB_CV405 Opened" : Real = PLC "PGC Flush_DB"."CV405 Opened", 1 s
   "PGC Flush_DB_CV401 Opened" : Bool = PLC "PGC Flush_DB"."CV401 Opened", 1 s
   "PGC Flush_DB_CV431 Opened" : Bool = PLC "PGC Flush_DB"."CV431 Opened", 1 s
   "PGC Flush_DB_CV403 Opened" : Real = PLC "PGC Flush_DB"."CV403 Opened", 1 s
   "PGC Flush_DB_CV441 Closed" : Bool = PLC "PGC Flush_DB"."CV441 Closed", 1 s
   "PGC Flush_DB_CAB Started" : Bool = PLC "PGC Flush_DB"."CAB Started", 1 s
   "50_CMND_DATA_CV403 Modulate Cmd" : Bool = PLC "50_CMND_DATA"."CV403 Modulate Cmd" AT %DB50.DBX6.0, 1 s
   "1403_PID_300CV403_State" : Int = PLC "1403_PID_300CV403".State, 1 s
   "PGC Flush_DB_PGC Stoped" : Bool = PLC "PGC Flush_DB"."PGC Stoped", 1 s
   "1405_PID_CV405_ManualValue" : Real = PLC "1405_PID_CV405".ManualValue, 1 s
   "1403_PID_300CV403_ModeActivate" : Bool = PLC "1403_PID_300CV403".ModeActivate, 1 s
   "1403_PID_300CV403_ManualEnable" : Bool = PLC "1403_PID_300CV403".ManualEnable, 1 s
   "1405_PID_CV405_ManualEnable" : Bool = PLC "1405_PID_CV405".ManualEnable, 1 s
   "2062_Warning_Data_BTCS_WARNING_WORD_01" : Word = PLC "2062_Warning_Data".BTCS_WARNING_WORD_01 AT %DB2062.DBW0, 1 s
   "2062_Warning_Data_BTCS_WARNING_WORD_02" : Word = PLC "2062_Warning_Data".BTCS_WARNING_WORD_02 AT %DB2062.DBW2, 1 s
   "2062_Warning_Data_BTCS_WARNING_WORD_03" : Word = PLC "2062_Warning_Data".BTCS_WARNING_WORD_03 AT %DB2062.DBW4, 1 s
   "2062_Warning_Data_BTCS_WARNING_WORD_04" : Word = PLC "2062_Warning_Data".BTCS_WARNING_WORD_04 AT %DB2062.DBW6, 1 s
   "2062_Warning_Data_BTCS_WARNING_WORD_05" : Word = PLC "2062_Warning_Data".BTCS_WARNING_WORD_05 AT %DB2062.DBW8, 1 s
   "2062_Warning_Data_BTCS_WARNING_WORD_06" : Word = PLC "2062_Warning_Data".BTCS_WARNING_WORD_06 AT %DB2062.DBW10, 1 s
   "2062_Warning_Data_BTCS_WARNING_WORD_07" : Word = PLC "2062_Warning_Data".BTCS_WARNING_WORD_07 AT %DB2062.DBW12, 1 s
   "2062_Warning_Data_BTCS_WARNING_WORD_08" : Word = PLC "2062_Warning_Data".BTCS_WARNING_WORD_08 AT %DB2062.DBW14, 1 s
   "2062_Warning_Data_BTCS_WARNING_WORD_09" : Word = PLC "2062_Warning_Data".BTCS_WARNING_WORD_09 AT %DB2062.DBW16, 1 s
   "2062_Warning_Data_BTCS_WARNING_WORD_10" : Word = PLC "2062_Warning_Data".BTCS_WARNING_WORD_10 AT %DB2062.DBW18, 1 s
   "2062_Warning_Data_BTCS_WARNING_WORD_11" : Word = PLC "2062_Warning_Data".BTCS_WARNING_WORD_11 AT %DB2062.DBW20, 1 s
   "80_From_HMI_PGC_RST_HRS" : Bool = PLC "80_From_HMI".PGC_RST_HRS, 1 s
   "102_Pilot_Burner_DB_FD_VRFCTN_TMR_Q" : Bool = PLC "102_Pilot_Burner_DB".FD_VRFCTN_TMR.Q, 1 s
   "102_Pilot_Burner_DB_FD_VRFCTN_TMR_ET" : Time = PLC "102_Pilot_Burner_DB".FD_VRFCTN_TMR.ET, 1 s
   "102_Pilot_Burner_DB_FD_VRFCTN_TMR II_ET" : Time = PLC "102_Pilot_Burner_DB"."FD_VRFCTN_TMR II".ET, 1 s
   "86_Times_PIT358 Delay" : Time = PLC "86_Times"."PIT358 Delay", 1 s
   "86_Times_PIT348 Delay" : Time = PLC "86_Times"."PIT348 Delay", 1 s
   "PGC Flush_DB_Temperature Setpoint" : Real = PLC "PGC Flush_DB"."Temperature Setpoint", 1 s
   "2062_Warning_Data_Water Level Override" : Bool = PLC "2062_Warning_Data"."Water Level Override" AT %DB2062.DBX376.0, 1 s
   "2062_Warning_Data_Water Level Override_Aux" : Bool = PLC "2062_Warning_Data"."Water Level Override_Aux" AT %DB2062.DBX376.2, 1 s
   "Sequence Times_DB_Boost" : Bool = PLC "Sequence Times_DB".Boost, 1 s
   "86_Times_FS317 delay" : Time = PLC "86_Times"."FS317 delay", 1 s
   "86_Times_FS320 delay" : Time = PLC "86_Times"."FS320 delay", 1 s
   "86_Times_PS101 Alarm Delay" : Time = PLC "86_Times"."PS101 Alarm Delay", 1 s
   "82_To_HMI_FS350 Animation" : Int = PLC "82_To_HMI"."FS350 Animation", 1 s
   "E-400 Animation_DB_Animation" : Int = PLC "E-400 Animation_DB".Animation, 1 s
   "1405_PID_CV405_Progress" : Real = PLC "1405_PID_CV405".Progress, 1 s
   "P304 Animation_IDB_Animation" : Int = PLC "P304 Animation_IDB".Animation, 1 s
   "FS332 Animation_IDB_Animation" : Int = PLC "FS332 Animation_IDB".Animation, 1 s
   "51_SLAVE_STATUS_MAIN_BURNER_ACTV" : Bool = PLC "51_SLAVE_STATUS".MAIN_BURNER_ACTV AT %DB51.DBX17.5, 1 s
   "Main Burner Animation_DB_Animation" : Int = PLC "Main Burner Animation_DB".Animation, 1 s
   "Sequence Times_DB_Post-Dwell Timer_Q" : Bool = PLC "Sequence Times_DB"."Post-Dwell Timer".Q, 1 s
      on ChangeValue: "TreatmentCycleCompleted"()
   "20_TANKS_IP_DATA_RIO_01_FIRST_TANK_MBG_FLOW N" : Real = PLC "20_TANKS_IP_DATA".RIO_01.FIRST_TANK."MBG_FLOW N", 1 s
   "20_TANKS_IP_DATA_RIO_01_FIRST_TANK_USD FLOW  N" : Real = PLC "20_TANKS_IP_DATA".RIO_01.FIRST_TANK."USD FLOW  N", 1 s
   "20_TANKS_IP_DATA_RIO_01_SECOND_TANK_MBG_FLOW N" : Real = PLC "20_TANKS_IP_DATA".RIO_01.SECOND_TANK."MBG_FLOW N", 1 s
   "20_TANKS_IP_DATA_RIO_01_SECOND_TANK_USD FLOW  N" : Real = PLC "20_TANKS_IP_DATA".RIO_01.SECOND_TANK."USD FLOW  N", 1 s
   "20_TANKS_IP_DATA_RIO_01_THIRD_TANK_MBG_FLOW N" : Real = PLC "20_TANKS_IP_DATA".RIO_01.THIRD_TANK."MBG_FLOW N", 1 s
   "20_TANKS_IP_DATA_RIO_01_THIRD_TANK_USD FLOW  N" : Real = PLC "20_TANKS_IP_DATA".RIO_01.THIRD_TANK."USD FLOW  N", 1 s
   "20_TANKS_IP_DATA_RIO_02_FIRST_TANK_MBG_FLOW N" : Real = PLC "20_TANKS_IP_DATA".RIO_02.FIRST_TANK."MBG_FLOW N" AT %DB1.DBD0, 1 s
   "20_TANKS_IP_DATA_RIO_02_FIRST_TANK_USD FLOW  N" : Real = PLC "20_TANKS_IP_DATA".RIO_02.FIRST_TANK."USD FLOW  N" AT %DB1.DBD0, 1 s
   "20_TANKS_IP_DATA_RIO_02_SECOND_TANK_MBG_FLOW N" : Real = PLC "20_TANKS_IP_DATA".RIO_02.SECOND_TANK."MBG_FLOW N" AT %DB1.DBD0, 1 s
   "20_TANKS_IP_DATA_RIO_02_SECOND_TANK_USD FLOW  N" : Real = PLC "20_TANKS_IP_DATA".RIO_02.SECOND_TANK."USD FLOW  N" AT %DB1.DBD0, 1 s
   "20_TANKS_IP_DATA_RIO_03_FIRST_TANK_MBG_FLOW N" : Real = PLC "20_TANKS_IP_DATA".RIO_03.FIRST_TANK."MBG_FLOW N", 1 s
   "20_TANKS_IP_DATA_RIO_03_FIRST_TANK_USD FLOW  N" : Real = PLC "20_TANKS_IP_DATA".RIO_03.FIRST_TANK."USD FLOW  N", 1 s
   "20_TANKS_IP_DATA_RIO_03_SECOND_TANK_MBG_FLOW N" : Real = PLC "20_TANKS_IP_DATA".RIO_03.SECOND_TANK."MBG_FLOW N", 1 s
   "20_TANKS_IP_DATA_RIO_03_SECOND_TANK_USD FLOW  N" : Real = PLC "20_TANKS_IP_DATA".RIO_03.SECOND_TANK."USD FLOW  N", 1 s
   "20_TANKS_IP_DATA_RIO_04_FIRST_TANK_MBG_FLOW N" : Real = PLC "20_TANKS_IP_DATA".RIO_04.FIRST_TANK."MBG_FLOW N", 1 s
   "20_TANKS_IP_DATA_RIO_04_FIRST_TANK_USD FLOW  N" : Real = PLC "20_TANKS_IP_DATA".RIO_04.FIRST_TANK."USD FLOW  N", 1 s
   "20_TANKS_IP_DATA_RIO_04_SECOND_TANK_MBG_FLOW N" : Real = PLC "20_TANKS_IP_DATA".RIO_04.SECOND_TANK."MBG_FLOW N", 1 s
   "20_TANKS_IP_DATA_RIO_04_SECOND_TANK_USD FLOW  N" : Real = PLC "20_TANKS_IP_DATA".RIO_04.SECOND_TANK."USD FLOW  N", 1 s
   "20_TANKS_IP_DATA_RIO_05_FIRST_TANK_MBG_FLOW N" : Real = PLC "20_TANKS_IP_DATA".RIO_05.FIRST_TANK."MBG_FLOW N", 1 s
   "20_TANKS_IP_DATA_RIO_05_FIRST_TANK_USD FLOW  N" : Real = PLC "20_TANKS_IP_DATA".RIO_05.FIRST_TANK."USD FLOW  N", 1 s
   "20_TANKS_IP_DATA_RIO_05_SECOND_TANK_USD FLOW  N" : Real = PLC "20_TANKS_IP_DATA".RIO_05.SECOND_TANK."USD FLOW  N", 1 s
   "20_TANKS_IP_DATA_RIO_06_FIRST_TANK_MBG_FLOW N" : Real = PLC "20_TANKS_IP_DATA".RIO_06.FIRST_TANK."MBG_FLOW N", 1 s
   "20_TANKS_IP_DATA_RIO_06_FIRST_TANK_USD FLOW  N" : Real = PLC "20_TANKS_IP_DATA".RIO_06.FIRST_TANK."USD FLOW  N", 1 s
   "20_TANKS_IP_DATA_RIO_06_SECOND_TANK_MBG_FLOW N" : Real = PLC "20_TANKS_IP_DATA".RIO_06.SECOND_TANK."MBG_FLOW N", 1 s
   "20_TANKS_IP_DATA_RIO_06_SECOND_TANK_USD FLOW  N" : Real = PLC "20_TANKS_IP_DATA".RIO_06.SECOND_TANK."USD FLOW  N", 1 s
   "20_TANKS_IP_DATA_RIO_07_FIRST_TANK_MBG_FLOW N" : Real = PLC "20_TANKS_IP_DATA".RIO_07.FIRST_TANK."MBG_FLOW N", 1 s
   "20_TANKS_IP_DATA_RIO_07_FIRST_TANK_USD FLOW  N" : Real = PLC "20_TANKS_IP_DATA".RIO_07.FIRST_TANK."USD FLOW  N", 1 s
   "Nm³/hr to m³/hr" : Bool = PLC "80_From_HMI"."m³/hr to Nm³/hr" AT %DB1.DBX0.0, 1 s
   "20_TANKS_IP_DATA_RIO_05_SECOND_TANK_MBG_FLOW N" : Real = PLC "20_TANKS_IP_DATA".RIO_05.SECOND_TANK."MBG_FLOW N", 1 s
   "IDB_E500A_Animation_Animation" : Int = PLC IDB_E500A_Animation.Animation, 1 s
   "IDB_E500B_Animation_Animation" : Int = PLC IDB_E500B_Animation.Animation, 1 s
   "Ful Pump Ani Animation_DB_Animation" : Int = PLC "Ful Pump Ani Animation_DB".Animation, 1 s
   "IDB_E131_Animation_Animation" : Int = PLC IDB_E131_Animation.Animation, 1 s
   "2062_Warning_Data_BTCS_WARNING_WORD_17" : Word = PLC "2062_Warning_Data".BTCS_WARNING_WORD_17 AT %DB2062.DBW372, 1 s
   "CCR HMI HEART BEAT" : Bool = PLC "59_COMMS_HEALTH_DATA"."CCR HMI HB" AT %DB1.DBX0.0, 100 ms
   "TRUE" : Bool = PLC AlwaysTRUE AT %M1.2, 1 s
   "IGG PLC HEART BEAT" : Bool = PLC "55_STATUS_DATA".HEART_BEAT AT %DB55.DBX0.0, 100 ms
      on ChangeValue: "HeartBeatFunction"()
   "80_From_HMI_Jurney Start Simulator" : Bool = PLC "80_From_HMI"."Jurney Start Simulator", 1 s
   "68_Sys_Status_Data_LOG IGG Simulator" : Bool = PLC "68_Sys_Status_Data"."LOG IGG Simulator", 1 s
   "68_Sys_Status_Data_LOG GCU Simulator" : Bool = PLC "68_Sys_Status_Data"."LOG GCU Simulator", 1 s
   "Setpoint Override_DB_Pressure Struct_Pressure Safe Set" : Real = PLC "Setpoint Override_DB"."Pressure Safe Target", 1 s
   "Setpoint Override_DB_Activate Temp Prot" : Bool = PLC "Setpoint Override_DB"."Activate Temp Prot", 1 s
   "Setpoint Override_DB_Activate Press Prot" : Bool = PLC "Setpoint Override_DB"."Activate Press Prot", 1 s
   "Setpoint Override_DB_Temperature Tolerance" : Real = PLC "Setpoint Override_DB"."Temperature Tolerance", 1 s
   "Setpoint Override_DB_Pressure Tolerance" : Real = PLC "Setpoint Override_DB"."Pressure Tolerance", 1 s
   "Setpoint Override_DB_Tank Change TimeOut" : Time = PLC "Setpoint Override_DB"."Tank Change TimeOut", 1 s
   "Setpoint Override_DB_Reset" : Bool = PLC "Setpoint Override_DB".Reset, 1 s
   "Setpoint Override_DB_Set Pressure" : Bool = PLC "Setpoint Override_DB"."Set Pressure", 1 s
      on ChangeValue: function_efd93a16("PGC Protection Warning", 300, 200, -1, 3, 1)
   "80_From_HMI_TT002 Target Protection" : Bool = PLC "80_From_HMI"."TT002 Target Protection", 1 s
   "80_From_HMI_PT002 Target Protection" : Bool = PLC "80_From_HMI"."PT002 Target Protection", 1 s
   "80_From_HMI_Tank Close Protection" : Bool = PLC "80_From_HMI"."Tank Close Protection", 1 s
   "84_Setpoints_PIT416_Target_Safe" : Real = PLC "84_Setpoints".PIT416_Target_Safe, 1 s
   "84_Setpoints_Tank Close TimeOut" : Time = PLC "84_Setpoints"."Tank Close TimeOut", 1 s
   "84_Setpoints_E-400 PT002 Tolerance" : Real = PLC "84_Setpoints"."E-400 PT002 Tolerance", 1 s
   "84_Setpoints_E-400 TT002 Tolerance" : Real = PLC "84_Setpoints"."E-400 TT002 Tolerance", 1 s
   "Sequence Times_DB_Jurney Timer_Days Left" : DInt = PLC "Sequence Times_DB"."Jurney Timer"."Days Left", 1 s
   "Sequence Times_DB_Jurney Timer_Hours Left" : DInt = PLC "Sequence Times_DB"."Jurney Timer"."Hours Left", 1 s
   "Sequence Times_DB_Jurney Timer_Minutes Left" : DInt = PLC "Sequence Times_DB"."Jurney Timer"."Minutes Left", 1 s
   "Warn To Start IGG-Last" : Bool = PLC "82_To_HMI"."Warn to Start IGG-Last", 1 s
      on ChangeValue: "TreatmentRequired"()
   "Warn To Start GCU" : Bool = PLC "82_To_HMI"."Warn to Start GCU", 1 s
      on ChangeValue: "TimeRemainingToRe_Ox"()
   "Warn To Start GCU-Last" : Bool = PLC "82_To_HMI"."Warn to Start GCU-Last", 1 s
      on ChangeValue: "TreatmentRequired_GCU"()
   "2086_Times_Stage Warning" : Time = PLC "2086_Times"."Stage Warning", 1 s
   "80_From_HMI_GCU Start Confirmed" : Bool = PLC "80_From_HMI"."GCU Start Confirmed", 1 s
   "102_Pilot_Burner_DB_STATE" : Int = PLC "102_Pilot_Burner_DB".STATE, 1 s
   "2068_Sys_Status_Data_Times Visibil" : Bool = PLC "2068_Sys_Status_Data"."Times Visibil", 1 s
   "Sequence Times_DB_Warn to GCU Start" : Bool = PLC "Sequence Times_DB"."Warn to GCU Start", 1 s
   "80_From_HMI_CSW OVR Stop" : Bool = PLC "80_From_HMI"."CSW OVR Stop", 1 s
   "Sequence Times_DB_Offset Timer_Days Left" : DInt = PLC "Sequence Times_DB"."Offset Timer"."Days Left", 1 s
   "Sequence Times_DB_Offset Timer_Hours Left" : DInt = PLC "Sequence Times_DB"."Offset Timer"."Hours Left", 1 s
   "Sequence Times_DB_Offset Timer_Minutes Left" : DInt = PLC "Sequence Times_DB"."Offset Timer"."Minutes Left", 1 s
   "Voyage Time Invalid" : Bool = PLC "Sequence Times_DB"."Voiage Time Invalid" AT %DB1.DBX0.0, 1 s
      on ChangeValue: "VoyageTimeInsufficient"()
   "82_To_HMI_IGG RUN Indication" : Bool = PLC "82_To_HMI"."IGG RUN Indication", 1 s
   "Not TANK Activ Warning" : Bool = PLC "2068_Sys_Status_Data"."Not TANK Activ Warning" AT %DB1.DBX0.0, 1 s
      on ChangeValue: "TANK_Activ_Warning"()
   "Sequence Times_DB_Pre-Dwell Done" : Bool = PLC "Sequence Times_DB"."Pre-Dwell Done", 1 s
   "Sequence Times_DB_De-Ox Done" : Bool = PLC "Sequence Times_DB"."De-Ox Done", 1 s
   "Sequence Times_DB_Dwell Done" : Bool = PLC "Sequence Times_DB"."Dwell Done", 1 s
   "Sequence Times_DB_Re-Ox Done" : Bool = PLC "Sequence Times_DB"."Re-Ox Done", 1 s
   "Sequence Times_DB_Post-Dwell Done" : Bool = PLC "Sequence Times_DB"."Post-Dwell Done", 1 s

HMI tags "Alarms"
   "60_Alarm_Data_BC_ALARM_WORD_01" : Word = PLC "60_Alarm_Data".BC_ALARM_WORD_01 AT %DB60.DBW0, 1 s
   "60_Alarm_Data_BC_ALARM_WORD_02" : Word = PLC "60_Alarm_Data".BC_ALARM_WORD_02 AT %DB60.DBW2, 1 s
   "60_Alarm_Data_BC_ALARM_WORD_03" : Word = PLC "60_Alarm_Data".BC_ALARM_WORD_03 AT %DB60.DBW4, 1 s
   "60_Alarm_Data_BC_ALARM_WORD_04" : Word = PLC "60_Alarm_Data".BC_ALARM_WORD_04 AT %DB60.DBW6, 1 s
   "60_Alarm_Data_IGG_ALARM_WORD_01" : Word = PLC "60_Alarm_Data".IGG_ALARM_WORD_01 AT %DB60.DBW0, 1 s
   "60_Alarm_Data_IGG_ALARM_WORD_02" : Word = PLC "60_Alarm_Data".IGG_ALARM_WORD_02 AT %DB60.DBW2, 1 s
   "60_Alarm_Data_IGG_ALARM_WORD_03" : Word = PLC "60_Alarm_Data".IGG_ALARM_WORD_03 AT %DB60.DBW4, 1 s
   "60_Alarm_Data_IGG_ALARM_WORD_04" : Word = PLC "60_Alarm_Data".IGG_ALARM_WORD_04 AT %DB60.DBW6, 1 s

